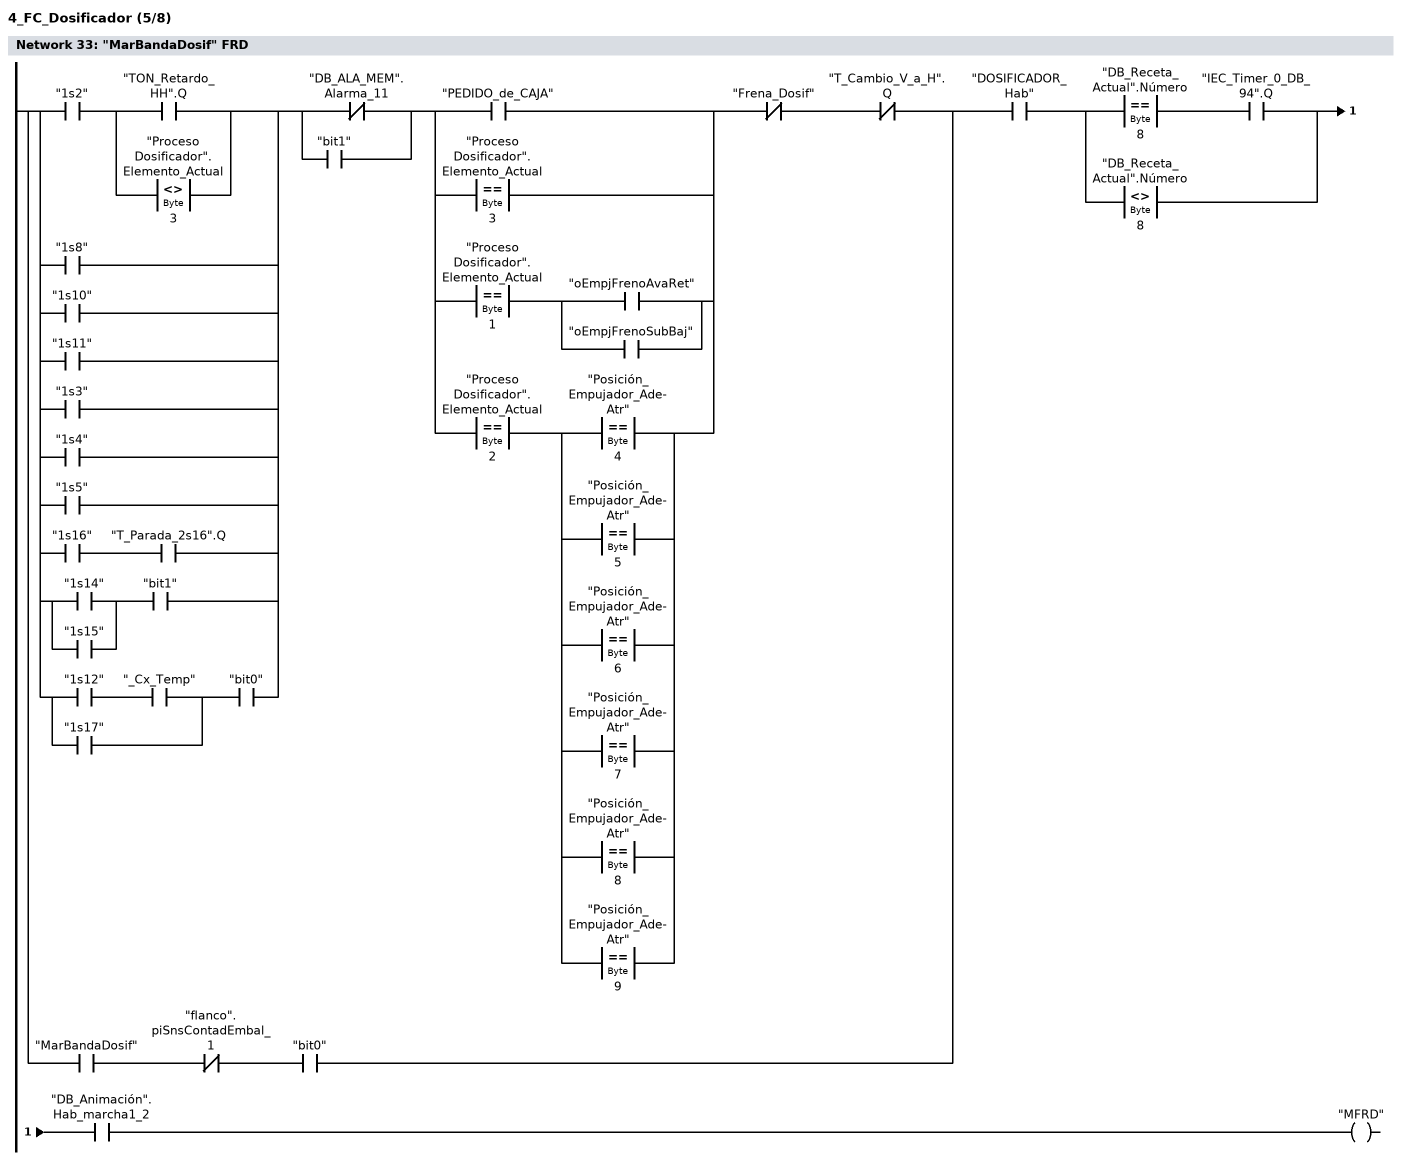
   RUNG wire#powerrail
      Contact( "1s2" )
      wire#w1
      Contact( "TON_Retardo_HH".Q )
      wire#w2
      I_Contact( "DB_ALA_MEM".Alarma_11 )
      wire#w5
      Contact( "PEDIDO_de_CAJA" )
      wire#w6
      I_Contact( "Frena_Dosif" )
      I_Contact( "T_Cambio_V_a_H".Q )
      wire#w9
      Contact( "DOSIFICADOR_Hab" )
      wire#w10
      { S7_Templates := "SrcType := Byte" } EQ_Contact(in1 := "DB_Receta_Actual".Número, in2 := 8)
      Contact( "IEC_Timer_0_DB_94".Q )
      wire#w11
      Contact( "DB_Animación".Hab_marcha1_2 )
      Coil( "MFRD" )
   END_RUNG
   RUNG wire#w1
      { S7_Templates := "SrcType := Byte" } NE_Contact(in1 := "Proceso Dosificador".Elemento_Actual, in2 := 3)
   END_RUNG wire#w2
   RUNG wire#powerrail
      Contact( "1s8" )
   END_RUNG wire#w2
   RUNG wire#powerrail
      Contact( "1s10" )
   END_RUNG wire#w2
   RUNG wire#powerrail
      Contact( "1s11" )
   END_RUNG wire#w2
   RUNG wire#powerrail
      Contact( "1s3" )
   END_RUNG wire#w2
   RUNG wire#powerrail
      Contact( "1s4" )
   END_RUNG wire#w2
   RUNG wire#powerrail
      Contact( "1s5" )
   END_RUNG wire#w2
   RUNG wire#powerrail
      Contact( "1s16" )
      Contact( "T_Parada_2s16".Q )
   END_RUNG wire#w2
   RUNG wire#powerrail
      Contact( "1s14" )
      wire#w3
      Contact( "bit1" )
   END_RUNG wire#w2
   RUNG wire#powerrail
      Contact( "1s15" )
   END_RUNG wire#w3
   RUNG wire#powerrail
      Contact( "1s12" )
      Contact( "_Cx_Temp" )
      wire#w4
      Contact( "bit0" )
   END_RUNG wire#w2
   RUNG wire#powerrail
      Contact( "1s17" )
   END_RUNG wire#w4
   RUNG wire#w2
      Contact( "bit1" )
   END_RUNG wire#w5
   RUNG wire#w5
      { S7_Templates := "SrcType := Byte" } EQ_Contact(in1 := "Proceso Dosificador".Elemento_Actual, in2 := 3)
   END_RUNG wire#w6
   RUNG wire#w5
      { S7_Templates := "SrcType := Byte" } EQ_Contact(in1 := "Proceso Dosificador".Elemento_Actual, in2 := 1)
      wire#w7
      Contact( "oEmpjFrenoAvaRet" )
   END_RUNG wire#w6
   RUNG wire#w7
      Contact( "oEmpjFrenoSubBaj" )
   END_RUNG wire#w6
   RUNG wire#w5
      { S7_Templates := "SrcType := Byte" } EQ_Contact(in1 := "Proceso Dosificador".Elemento_Actual, in2 := 2)
      wire#w8
      { S7_Templates := "SrcType := Byte" } EQ_Contact(in1 := "Posición_Empujador_Ade-Atr", in2 := 4)
   END_RUNG wire#w6
   RUNG wire#w8
      { S7_Templates := "SrcType := Byte" } EQ_Contact(in1 := "Posición_Empujador_Ade-Atr", in2 := 5)
   END_RUNG wire#w6
   RUNG wire#w8
      { S7_Templates := "SrcType := Byte" } EQ_Contact(in1 := "Posición_Empujador_Ade-Atr", in2 := 6)
   END_RUNG wire#w6
   RUNG wire#w8
      { S7_Templates := "SrcType := Byte" } EQ_Contact(in1 := "Posición_Empujador_Ade-Atr", in2 := 7)
   END_RUNG wire#w6
   RUNG wire#w8
      { S7_Templates := "SrcType := Byte" } EQ_Contact(in1 := "Posición_Empujador_Ade-Atr", in2 := 8)
   END_RUNG wire#w6
   RUNG wire#w8
      { S7_Templates := "SrcType := Byte" } EQ_Contact(in1 := "Posición_Empujador_Ade-Atr", in2 := 9)
   END_RUNG wire#w6
   RUNG wire#powerrail
      Contact( "MarBandaDosif" )
      I_Contact( "flanco".piSnsContadEmbal_1 )
      Contact( "bit0" )
   END_RUNG wire#w9
   RUNG wire#w10
      { S7_Templates := "SrcType := Byte" } NE_Contact(in1 := "DB_Receta_Actual".Número, in2 := 8)
   END_RUNG wire#w11
   // the same network as SCL:
   "MFRD" := (((("1s2" AND ("TON_Retardo_HH".Q OR ("Proceso Dosificador".Elemento_Actual <> 3))) OR "1s8" OR "1s10" OR "1s11" OR "1s3" OR "1s4" OR "1s5" OR ("1s16" AND "T_Parada_2s16".Q) OR (("1s14" OR "1s15") AND "bit1") OR ((("1s12" AND "_Cx_Temp") OR "1s17") AND "bit0")) AND (NOT "DB_ALA_MEM".Alarma_11 OR "bit1") AND ("PEDIDO_de_CAJA" OR ("Proceso Dosificador".Elemento_Actual = 3) OR (("Proceso Dosificador".Elemento_Actual = 1) AND ("oEmpjFrenoAvaRet" OR "oEmpjFrenoSubBaj")) OR (("Proceso Dosificador".Elemento_Actual = 2) AND (("Posición_Empujador_Ade-Atr" = 4) OR ("Posición_Empujador_Ade-Atr" = 5) OR ("Posición_Empujador_Ade-Atr" = 6) OR ("Posición_Empujador_Ade-Atr" = 7) OR ("Posición_Empujador_Ade-Atr" = 8) OR ("Posición_Empujador_Ade-Atr" = 9)))) AND NOT "Frena_Dosif" AND NOT "T_Cambio_V_a_H".Q) OR ("MarBandaDosif" AND NOT "flanco".piSnsContadEmbal_1 AND "bit0")) AND "DOSIFICADOR_Hab" AND ((("DB_Receta_Actual".Número = 8) AND "IEC_Timer_0_DB_94".Q) OR ("DB_Receta_Actual".Número <> 8)) AND "DB_Animación".Hab_marcha1_2;
END_REGION

REGION Network 34: "MarBandaDosif" IGS/CRJ
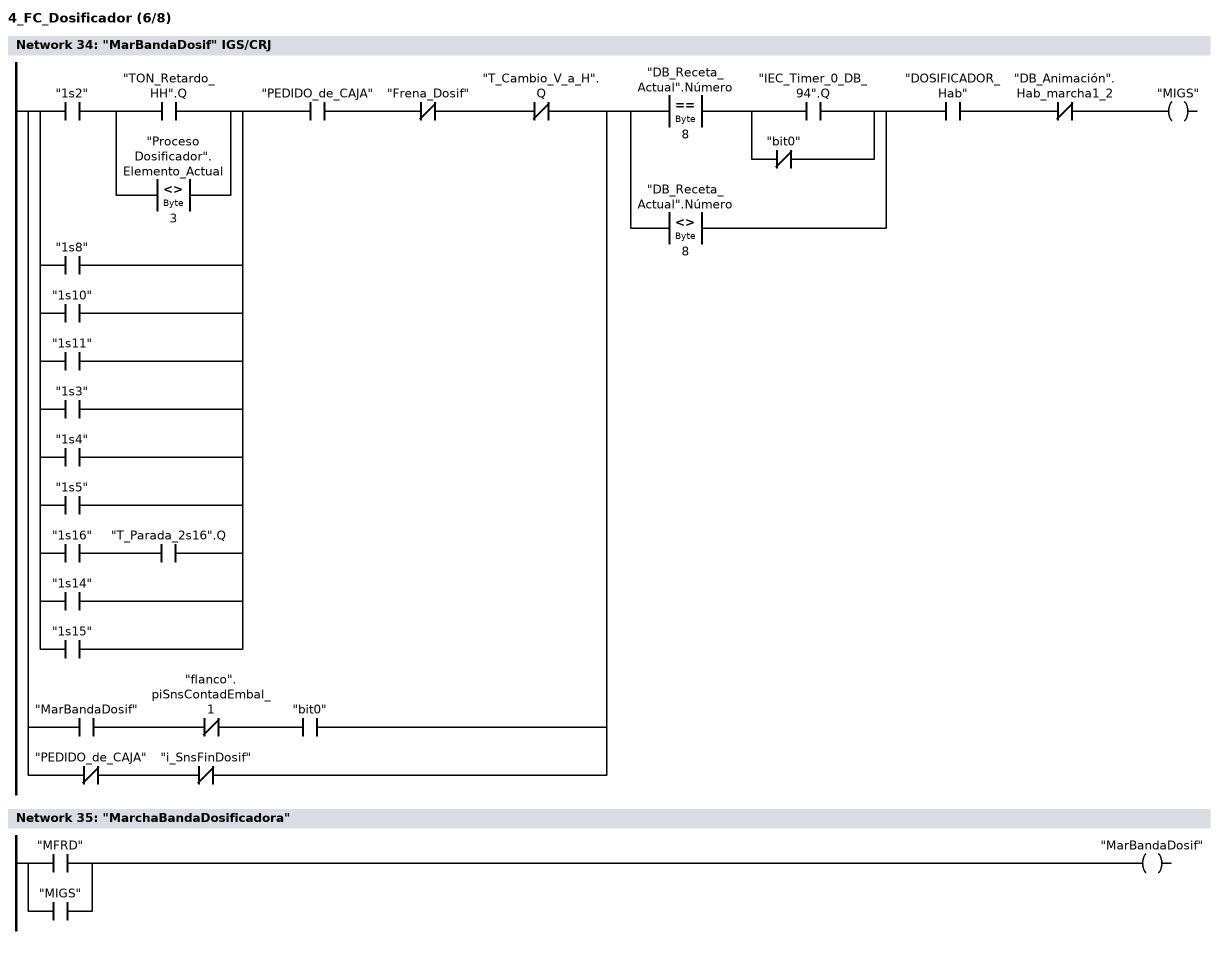
   RUNG wire#powerrail
      Contact( "1s2" )
      wire#w1
      Contact( "TON_Retardo_HH".Q )
      wire#w2
      Contact( "PEDIDO_de_CAJA" )
      I_Contact( "Frena_Dosif" )
      I_Contact( "T_Cambio_V_a_H".Q )
      wire#w3
      { S7_Templates := "SrcType := Byte" } EQ_Contact(in1 := "DB_Receta_Actual".Número, in2 := 8)
      wire#w4
      Contact( "IEC_Timer_0_DB_94".Q )
      wire#w5
      Contact( "DOSIFICADOR_Hab" )
      I_Contact( "DB_Animación".Hab_marcha1_2 )
      Coil( "MIGS" )
   END_RUNG
   RUNG wire#w1
      { S7_Templates := "SrcType := Byte" } NE_Contact(in1 := "Proceso Dosificador".Elemento_Actual, in2 := 3)
   END_RUNG wire#w2
   RUNG wire#powerrail
      Contact( "1s8" )
   END_RUNG wire#w2
   RUNG wire#powerrail
      Contact( "1s10" )
   END_RUNG wire#w2
   RUNG wire#powerrail
      Contact( "1s11" )
   END_RUNG wire#w2
   RUNG wire#powerrail
      Contact( "1s3" )
   END_RUNG wire#w2
   RUNG wire#powerrail
      Contact( "1s4" )
   END_RUNG wire#w2
   RUNG wire#powerrail
      Contact( "1s5" )
   END_RUNG wire#w2
   RUNG wire#powerrail
      Contact( "1s16" )
      Contact( "T_Parada_2s16".Q )
   END_RUNG wire#w2
   RUNG wire#powerrail
      Contact( "1s14" )
   END_RUNG wire#w2
   RUNG wire#powerrail
      Contact( "1s15" )
   END_RUNG wire#w2
   RUNG wire#powerrail
      Contact( "MarBandaDosif" )
      I_Contact( "flanco".piSnsContadEmbal_1 )
      Contact( "bit0" )
   END_RUNG wire#w3
   RUNG wire#powerrail
      I_Contact( "PEDIDO_de_CAJA" )
      I_Contact( "i_SnsFinDosif" )
   END_RUNG wire#w3
   RUNG wire#w4
      I_Contact( "bit0" )
   END_RUNG wire#w5
   RUNG wire#w3
      { S7_Templates := "SrcType := Byte" } NE_Contact(in1 := "DB_Receta_Actual".Número, in2 := 8)
   END_RUNG wire#w5
   // the same network as SCL:
   "MIGS" := (((("1s2" AND ("TON_Retardo_HH".Q OR ("Proceso Dosificador".Elemento_Actual <> 3))) OR "1s8" OR "1s10" OR "1s11" OR "1s3" OR "1s4" OR "1s5" OR ("1s16" AND "T_Parada_2s16".Q) OR "1s14" OR "1s15") AND "PEDIDO_de_CAJA" AND NOT "Frena_Dosif" AND NOT "T_Cambio_V_a_H".Q) OR ("MarBandaDosif" AND NOT "flanco".piSnsContadEmbal_1 AND "bit0") OR (NOT "PEDIDO_de_CAJA" AND NOT "i_SnsFinDosif")) AND ((("DB_Receta_Actual".Número = 8) AND ("IEC_Timer_0_DB_94".Q OR NOT "bit0")) OR ("DB_Receta_Actual".Número <> 8)) AND "DOSIFICADOR_Hab" AND NOT "DB_Animación".Hab_marcha1_2;
END_REGION

REGION Network 35: "MarchaBandaDosificadora"
   RUNG wire#powerrail
      Contact( "MFRD" )
      wire#w1
      Coil( "MarBandaDosif" )
   END_RUNG
   RUNG wire#powerrail
      Contact( "MIGS" )
   END_RUNG wire#w1
   // the same network as SCL:
   "MarBandaDosif" := "MFRD" OR "MIGS";
END_REGION

REGION Network 36: Temporizador provisario para Marcha Banda Dosifidicadora"
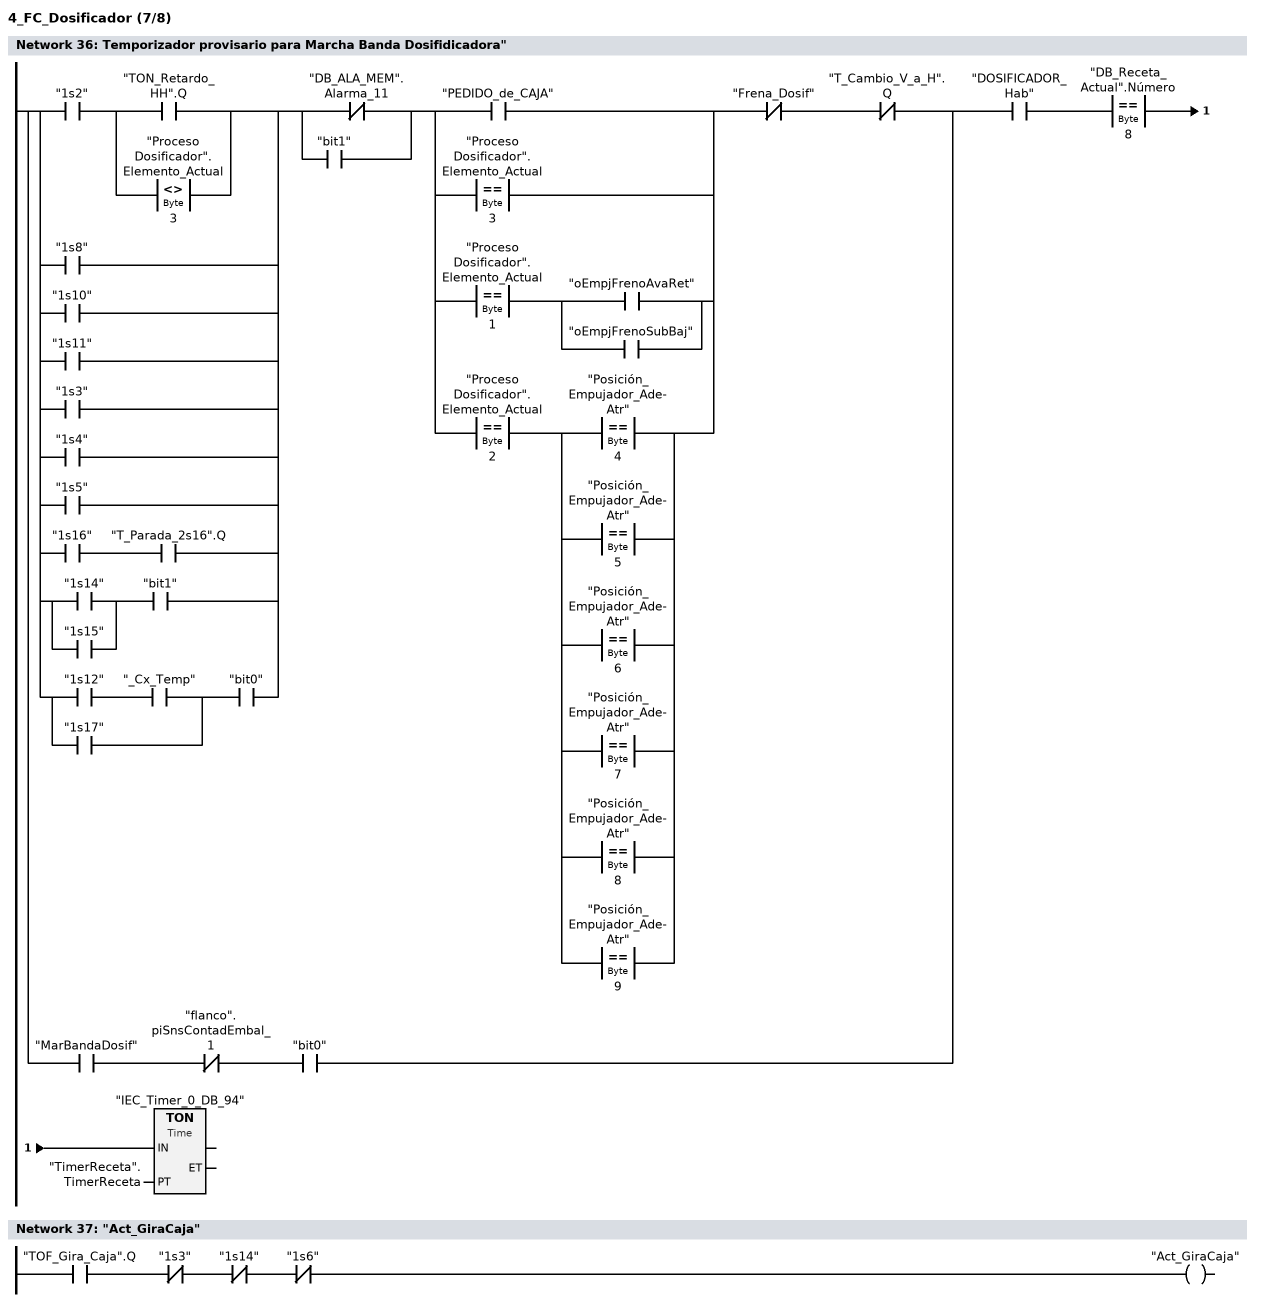
   "IEC_Timer_0_DB_94".TON(IN := (((("1s2" AND ("TON_Retardo_HH".Q OR ("Proceso Dosificador".Elemento_Actual <> 3))) OR "1s8" OR "1s10" OR "1s11" OR "1s3" OR "1s4" OR "1s5" OR ("1s16" AND "T_Parada_2s16".Q) OR (("1s14" OR "1s15") AND "bit1") OR ((("1s12" AND "_Cx_Temp") OR "1s17") AND "bit0")) AND (NOT "DB_ALA_MEM".Alarma_11 OR "bit1") AND ("PEDIDO_de_CAJA" OR ("Proceso Dosificador".Elemento_Actual = 3) OR (("Proceso Dosificador".Elemento_Actual = 1) AND ("oEmpjFrenoAvaRet" OR "oEmpjFrenoSubBaj")) OR (("Proceso Dosificador".Elemento_Actual = 2) AND (("Posición_Empujador_Ade-Atr" = 4) OR ("Posición_Empujador_Ade-Atr" = 5) OR ("Posición_Empujador_Ade-Atr" = 6) OR ("Posición_Empujador_Ade-Atr" = 7) OR ("Posición_Empujador_Ade-Atr" = 8) OR ("Posición_Empujador_Ade-Atr" = 9)))) AND NOT "Frena_Dosif" AND NOT "T_Cambio_V_a_H".Q) OR ("MarBandaDosif" AND NOT "flanco".piSnsContadEmbal_1 AND "bit0")) AND "DOSIFICADOR_Hab" AND ("DB_Receta_Actual".Número = 8),
                           PT := "TimerReceta".TimerReceta);
END_REGION

REGION Network 37: "Act_GiraCaja"
   RUNG wire#powerrail
      Contact( "TOF_Gira_Caja".Q )
      I_Contact( "1s3" )
      I_Contact( "1s14" )
      I_Contact( "1s6" )
      Coil( "Act_GiraCaja" )
   END_RUNG
   // the same network as SCL:
   "Act_GiraCaja" := "TOF_Gira_Caja".Q AND NOT "1s3" AND NOT "1s14" AND NOT "1s6";
END_REGION

REGION Network 38: "Act_EmpujaCaja"
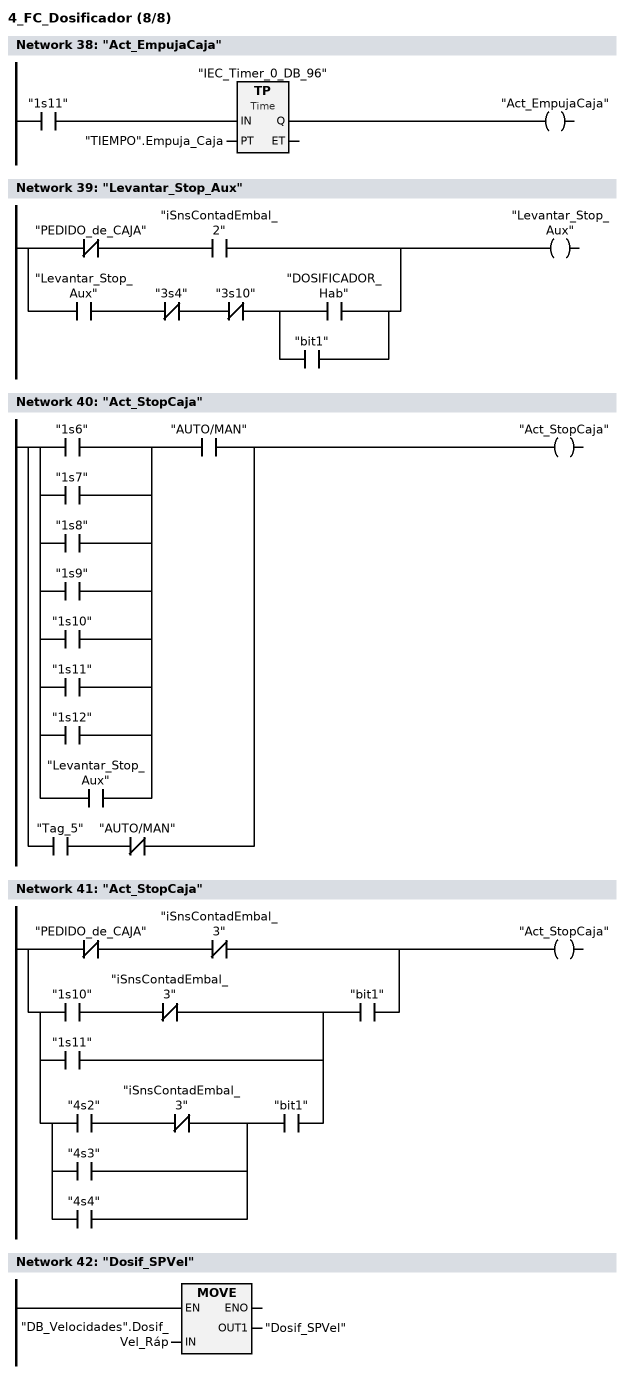
   "IEC_Timer_0_DB_96".TP(in := "1s11", pt := "TIEMPO".Empuja_Caja);
   "Act_EmpujaCaja" := "IEC_Timer_0_DB_96".q;
END_REGION

REGION Network 39: "Levantar_Stop_Aux"
   RUNG wire#powerrail
      I_Contact( "PEDIDO_de_CAJA" )
      Contact( "iSnsContadEmbal_2" )
      wire#w1
      Coil( "Levantar_Stop_Aux" )
   END_RUNG
   RUNG wire#powerrail
      Contact( "Levantar_Stop_Aux" )
      I_Contact( "3s4" )
      I_Contact( "3s10" )
      wire#w2
      Contact( "DOSIFICADOR_Hab" )
   END_RUNG wire#w1
   RUNG wire#w2
      Contact( "bit1" )
   END_RUNG wire#w1
   // the same network as SCL:
   "Levantar_Stop_Aux" := (NOT "PEDIDO_de_CAJA" AND "iSnsContadEmbal_2") OR ("Levantar_Stop_Aux" AND NOT "3s4" AND NOT "3s10" AND ("DOSIFICADOR_Hab" OR "bit1"));
END_REGION

REGION Network 40: "Act_StopCaja"
   RUNG wire#powerrail
      Contact( "1s6" )
      wire#w1
      Contact( "AUTO/MAN" )
      wire#w2
      Coil( "Act_StopCaja" )
   END_RUNG
   RUNG wire#powerrail
      Contact( "1s7" )
   END_RUNG wire#w1
   RUNG wire#powerrail
      Contact( "1s8" )
   END_RUNG wire#w1
   RUNG wire#powerrail
      Contact( "1s9" )
   END_RUNG wire#w1
   RUNG wire#powerrail
      Contact( "1s10" )
   END_RUNG wire#w1
   RUNG wire#powerrail
      Contact( "1s11" )
   END_RUNG wire#w1
   RUNG wire#powerrail
      Contact( "1s12" )
   END_RUNG wire#w1
   RUNG wire#powerrail
      Contact( "Levantar_Stop_Aux" )
   END_RUNG wire#w1
   RUNG wire#powerrail
      Contact( "Tag_5" )
      I_Contact( "AUTO/MAN" )
   END_RUNG wire#w2
   // the same network as SCL:
   "Act_StopCaja" := (("1s6" OR "1s7" OR "1s8" OR "1s9" OR "1s10" OR "1s11" OR "1s12" OR "Levantar_Stop_Aux") AND "AUTO/MAN") OR ("Tag_5" AND NOT "AUTO/MAN");
END_REGION

REGION Network 41: "Act_StopCaja"
   RUNG wire#powerrail
      I_Contact( "PEDIDO_de_CAJA" )
      I_Contact( "iSnsContadEmbal_3" )
      wire#w1
      Coil( "Act_StopCaja" )
   END_RUNG
   RUNG wire#powerrail
      Contact( "1s10" )
      I_Contact( "iSnsContadEmbal_3" )
      wire#w2
      Contact( "bit1" )
   END_RUNG wire#w1
   RUNG wire#powerrail
      Contact( "1s11" )
   END_RUNG wire#w2
   RUNG wire#powerrail
      Contact( "4s2" )
      I_Contact( "iSnsContadEmbal_3" )
      wire#w3
      Contact( "bit1" )
   END_RUNG wire#w2
   RUNG wire#powerrail
      Contact( "4s3" )
   END_RUNG wire#w3
   RUNG wire#powerrail
      Contact( "4s4" )
   END_RUNG wire#w3
   // the same network as SCL:
   "Act_StopCaja" := (NOT "PEDIDO_de_CAJA" AND NOT "iSnsContadEmbal_3") OR ((("1s10" AND NOT "iSnsContadEmbal_3") OR "1s11" OR ((("4s2" AND NOT "iSnsContadEmbal_3") OR "4s3" OR "4s4") AND "bit1")) AND "bit1");
END_REGION

REGION Network 42: "Dosif_SPVel"
   RUNG wire#powerrail
      { S7_GenerateENO := "TRUE" } Move(in := "DB_Velocidades".Dosif_Vel_Ráp, out1 => "Dosif_SPVel")
   END_RUNG
   // the same network as SCL:
   "Dosif_SPVel" := "DB_Velocidades".Dosif_Vel_Ráp;
END_REGION
END_FUNCTION

FUNCTION "5_FC_Empujador" : Void   // FC12, LAD
{ S7_Optimized_Access := 'FALSE' }
VERSION : 0.1
BEGIN

REGION Network 1
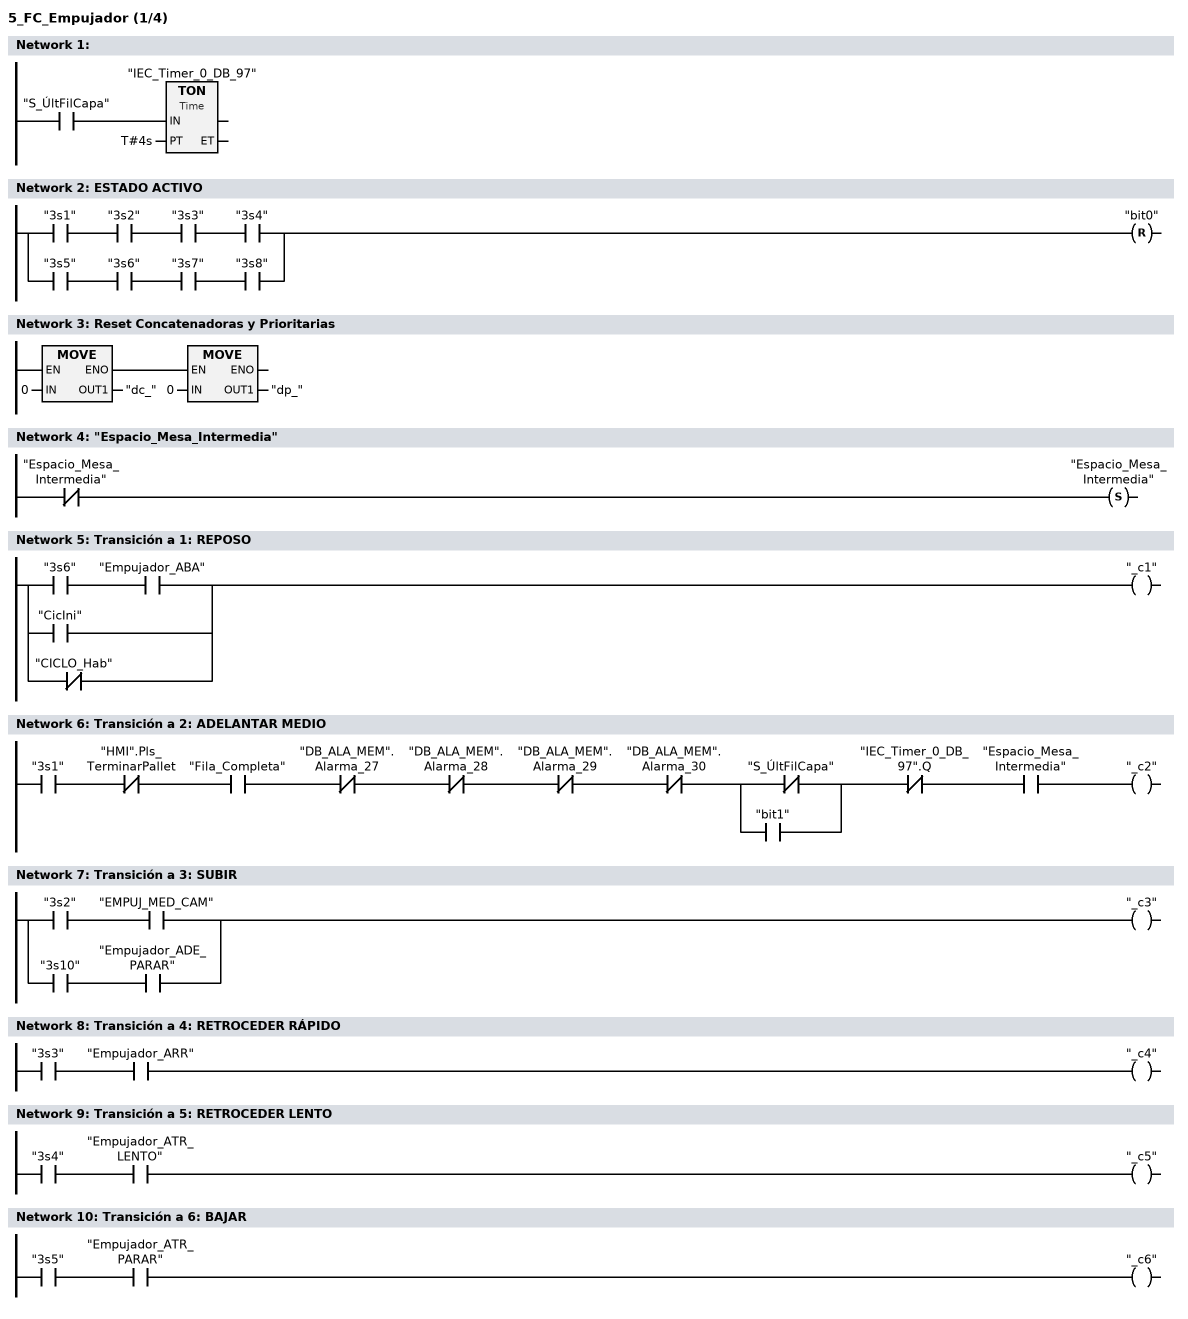
   "IEC_Timer_0_DB_97".TON(in := "S_ÚltFilCapa", pt := T#4s);
END_REGION

REGION Network 2: ESTADO ACTIVO
   RUNG wire#powerrail
      Contact( "3s1" )
      Contact( "3s2" )
      Contact( "3s3" )
      Contact( "3s4" )
      wire#w1
      R_Coil( "bit0" )
   END_RUNG
   RUNG wire#powerrail
      Contact( "3s5" )
      Contact( "3s6" )
      Contact( "3s7" )
      Contact( "3s8" )
   END_RUNG wire#w1
   // the same network as SCL:
   IF ("3s1" AND "3s2" AND "3s3" AND "3s4") OR ("3s5" AND "3s6" AND "3s7" AND "3s8") THEN
       "bit0" := FALSE;
   END_IF;
END_REGION

REGION Network 3: Reset Concatenadoras y Prioritarias
   RUNG wire#powerrail
      { S7_GenerateENO := "TRUE" } Move(in := 0, out1 => "dc_")
      { S7_GenerateENO := "TRUE" } Move(in := 0, out1 => "dp_")
   END_RUNG
   // the same network as SCL:
   // ENO of a box is taken as its EN; it also drops when the box reports an error
   "dc_" := 0;
   "dp_" := 0;
END_REGION

REGION Network 4: "Espacio_Mesa_Intermedia"
   RUNG wire#powerrail
      I_Contact( "Espacio_Mesa_Intermedia" )
      S_Coil( "Espacio_Mesa_Intermedia" )
   END_RUNG
   // the same network as SCL:
   IF NOT "Espacio_Mesa_Intermedia" THEN "Espacio_Mesa_Intermedia" := TRUE; END_IF;
END_REGION

REGION Network 5: Transición a 1: REPOSO
   RUNG wire#powerrail
      Contact( "3s6" )
      Contact( "Empujador_ABA" )
      wire#w1
      Coil( "_c1" )
   END_RUNG
   RUNG wire#powerrail
      Contact( "CicIni" )
   END_RUNG wire#w1
   RUNG wire#powerrail
      I_Contact( "CICLO_Hab" )
   END_RUNG wire#w1
   // the same network as SCL:
   "_c1" := ("3s6" AND "Empujador_ABA") OR "CicIni" OR NOT "CICLO_Hab";
END_REGION

REGION Network 6: Transición a 2: ADELANTAR MEDIO
   RUNG wire#powerrail
      Contact( "3s1" )
      I_Contact( "HMI".Pls_TerminarPallet )
      Contact( "Fila_Completa" )
      I_Contact( "DB_ALA_MEM".Alarma_27 )
      I_Contact( "DB_ALA_MEM".Alarma_28 )
      I_Contact( "DB_ALA_MEM".Alarma_29 )
      I_Contact( "DB_ALA_MEM".Alarma_30 )
      wire#w1
      I_Contact( "S_ÚltFilCapa" )
      wire#w2
      I_Contact( "IEC_Timer_0_DB_97".Q )
      Contact( "Espacio_Mesa_Intermedia" )
      Coil( "_c2" )
   END_RUNG
   RUNG wire#w1
      Contact( "bit1" )
   END_RUNG wire#w2
   // the same network as SCL:
   "_c2" := "3s1" AND NOT "HMI".Pls_TerminarPallet AND "Fila_Completa" AND NOT "DB_ALA_MEM".Alarma_27 AND NOT "DB_ALA_MEM".Alarma_28 AND NOT "DB_ALA_MEM".Alarma_29 AND NOT "DB_ALA_MEM".Alarma_30 AND (NOT "S_ÚltFilCapa" OR "bit1") AND NOT "IEC_Timer_0_DB_97".Q AND "Espacio_Mesa_Intermedia";
END_REGION

REGION Network 7: Transición a 3: SUBIR
   RUNG wire#powerrail
      Contact( "3s2" )
      Contact( "EMPUJ_MED_CAM" )
      wire#w1
      Coil( "_c3" )
   END_RUNG
   RUNG wire#powerrail
      Contact( "3s10" )
      Contact( "Empujador_ADE_PARAR" )
   END_RUNG wire#w1
   // the same network as SCL:
   "_c3" := ("3s2" AND "EMPUJ_MED_CAM") OR ("3s10" AND "Empujador_ADE_PARAR");
END_REGION

REGION Network 8: Transición a 4: RETROCEDER RÁPIDO
   RUNG wire#powerrail
      Contact( "3s3" )
      Contact( "Empujador_ARR" )
      Coil( "_c4" )
   END_RUNG
   // the same network as SCL:
   "_c4" := "3s3" AND "Empujador_ARR";
END_REGION

REGION Network 9: Transición a 5: RETROCEDER LENTO
   RUNG wire#powerrail
      Contact( "3s4" )
      Contact( "Empujador_ATR_LENTO" )
      Coil( "_c5" )
   END_RUNG
   // the same network as SCL:
   "_c5" := "3s4" AND "Empujador_ATR_LENTO";
END_REGION

REGION Network 10: Transición a 6: BAJAR
   RUNG wire#powerrail
      Contact( "3s5" )
      Contact( "Empujador_ATR_PARAR" )
      Coil( "_c6" )
   END_RUNG
   // the same network as SCL:
   "_c6" := "3s5" AND "Empujador_ATR_PARAR";
END_REGION

REGION Network 11: Transición a 7: ESPERAR PLATAFORMA
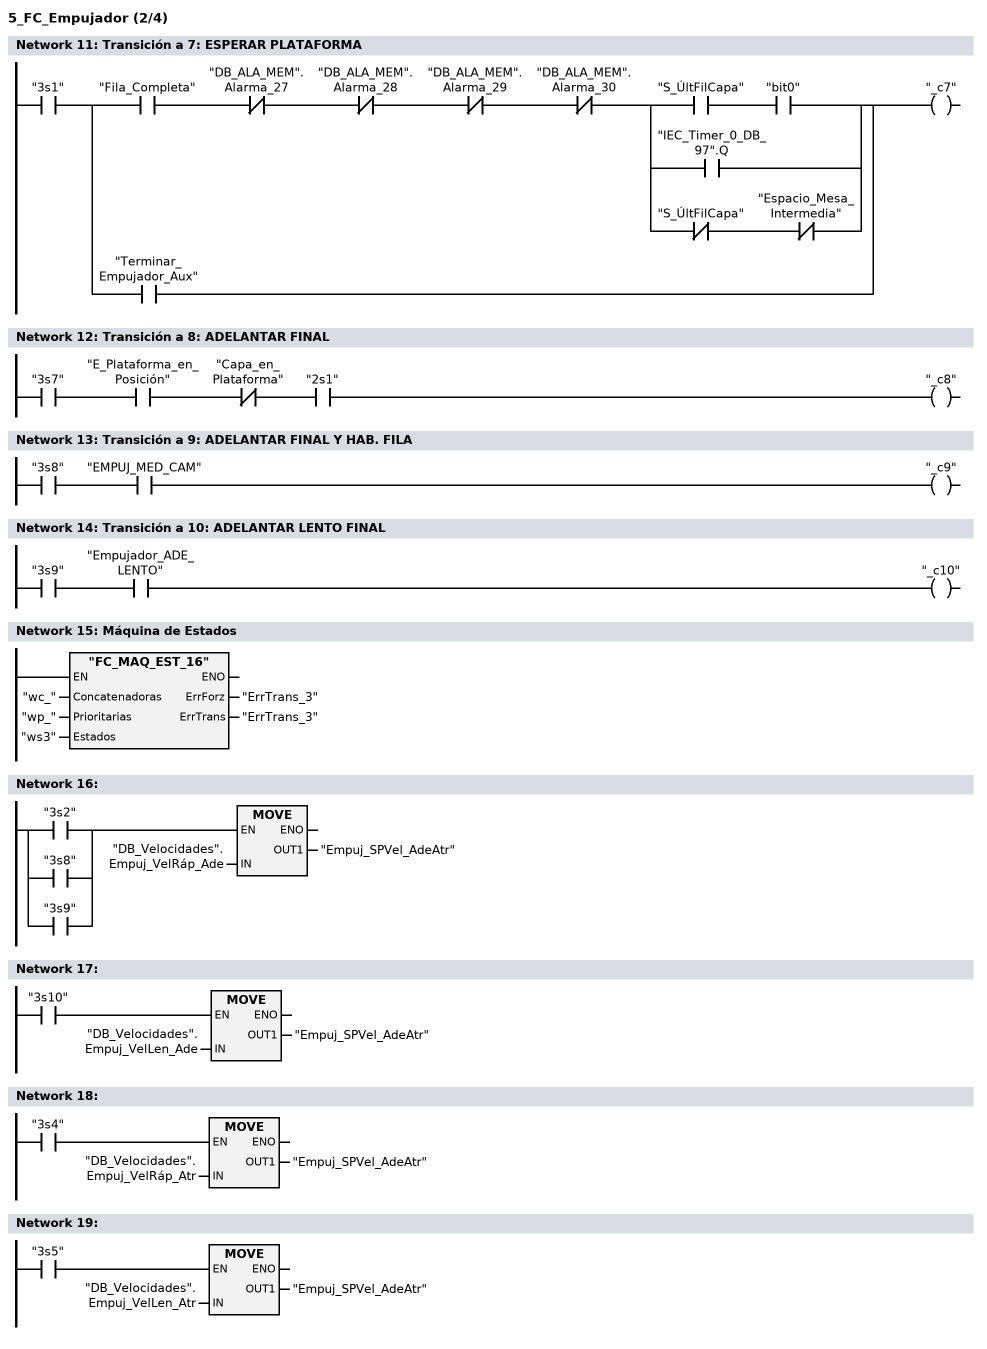
   RUNG wire#powerrail
      Contact( "3s1" )
      wire#w1
      Contact( "Fila_Completa" )
      I_Contact( "DB_ALA_MEM".Alarma_27 )
      I_Contact( "DB_ALA_MEM".Alarma_28 )
      I_Contact( "DB_ALA_MEM".Alarma_29 )
      I_Contact( "DB_ALA_MEM".Alarma_30 )
      wire#w2
      Contact( "S_ÚltFilCapa" )
      Contact( "bit0" )
      wire#w3
      Coil( "_c7" )
   END_RUNG
   RUNG wire#w2
      Contact( "IEC_Timer_0_DB_97".Q )
   END_RUNG wire#w3
   RUNG wire#w2
      I_Contact( "S_ÚltFilCapa" )
      I_Contact( "Espacio_Mesa_Intermedia" )
   END_RUNG wire#w3
   RUNG wire#w1
      Contact( "Terminar_Empujador_Aux" )
   END_RUNG wire#w3
   // the same network as SCL:
   "_c7" := "3s1" AND (("Fila_Completa" AND NOT "DB_ALA_MEM".Alarma_27 AND NOT "DB_ALA_MEM".Alarma_28 AND NOT "DB_ALA_MEM".Alarma_29 AND NOT "DB_ALA_MEM".Alarma_30 AND (("S_ÚltFilCapa" AND "bit0") OR "IEC_Timer_0_DB_97".Q OR (NOT "S_ÚltFilCapa" AND NOT "Espacio_Mesa_Intermedia"))) OR "Terminar_Empujador_Aux");
END_REGION

REGION Network 12: Transición a 8: ADELANTAR FINAL
   RUNG wire#powerrail
      Contact( "3s7" )
      Contact( "E_Plataforma_en_Posición" )
      I_Contact( "Capa_en_Plataforma" )
      Contact( "2s1" )
      Coil( "_c8" )
   END_RUNG
   // the same network as SCL:
   "_c8" := "3s7" AND "E_Plataforma_en_Posición" AND NOT "Capa_en_Plataforma" AND "2s1";
END_REGION

REGION Network 13: Transición a 9: ADELANTAR FINAL Y HAB. FILA
   RUNG wire#powerrail
      Contact( "3s8" )
      Contact( "EMPUJ_MED_CAM" )
      Coil( "_c9" )
   END_RUNG
   // the same network as SCL:
   "_c9" := "3s8" AND "EMPUJ_MED_CAM";
END_REGION

REGION Network 14: Transición a 10: ADELANTAR LENTO FINAL
   RUNG wire#powerrail
      Contact( "3s9" )
      Contact( "Empujador_ADE_LENTO" )
      Coil( "_c10" )
   END_RUNG
   // the same network as SCL:
   "_c10" := "3s9" AND "Empujador_ADE_LENTO";
END_REGION

REGION Network 15: Máquina de Estados
   RUNG wire#powerrail
      "FC_MAQ_EST_16"(Concatenadoras := "wc_", Prioritarias := "wp_", Estados := "ws3", ErrForz => "ErrTrans_3", ErrTrans => "ErrTrans_3")
   END_RUNG
   // the same network as SCL:
   "FC_MAQ_EST_16"(Concatenadoras := "wc_",
                   Prioritarias := "wp_",
                   Estados := "ws3",
                   ErrForz => "ErrTrans_3",
                   ErrTrans => "ErrTrans_3");
END_REGION

REGION Network 16
   RUNG wire#powerrail
      Contact( "3s2" )
      wire#w1
      { S7_GenerateENO := "TRUE" } Move(in := "DB_Velocidades".Empuj_VelRáp_Ade, out1 => "Empuj_SPVel_AdeAtr")
   END_RUNG
   RUNG wire#powerrail
      Contact( "3s8" )
   END_RUNG wire#w1
   RUNG wire#powerrail
      Contact( "3s9" )
   END_RUNG wire#w1
   // the same network as SCL:
   IF "3s2" OR "3s8" OR "3s9" THEN "Empuj_SPVel_AdeAtr" := "DB_Velocidades".Empuj_VelRáp_Ade; END_IF;
END_REGION

REGION Network 17
   RUNG wire#powerrail
      Contact( "3s10" )
      { S7_GenerateENO := "TRUE" } Move(in := "DB_Velocidades".Empuj_VelLen_Ade, out1 => "Empuj_SPVel_AdeAtr")
   END_RUNG
   // the same network as SCL:
   IF "3s10" THEN "Empuj_SPVel_AdeAtr" := "DB_Velocidades".Empuj_VelLen_Ade; END_IF;
END_REGION

REGION Network 18
   RUNG wire#powerrail
      Contact( "3s4" )
      { S7_GenerateENO := "TRUE" } Move(in := "DB_Velocidades".Empuj_VelRáp_Atr, out1 => "Empuj_SPVel_AdeAtr")
   END_RUNG
   // the same network as SCL:
   IF "3s4" THEN "Empuj_SPVel_AdeAtr" := "DB_Velocidades".Empuj_VelRáp_Atr; END_IF;
END_REGION

REGION Network 19
   RUNG wire#powerrail
      Contact( "3s5" )
      { S7_GenerateENO := "TRUE" } Move(in := "DB_Velocidades".Empuj_VelLen_Atr, out1 => "Empuj_SPVel_AdeAtr")
   END_RUNG
   // the same network as SCL:
   IF "3s5" THEN "Empuj_SPVel_AdeAtr" := "DB_Velocidades".Empuj_VelLen_Atr; END_IF;
END_REGION

REGION Network 20
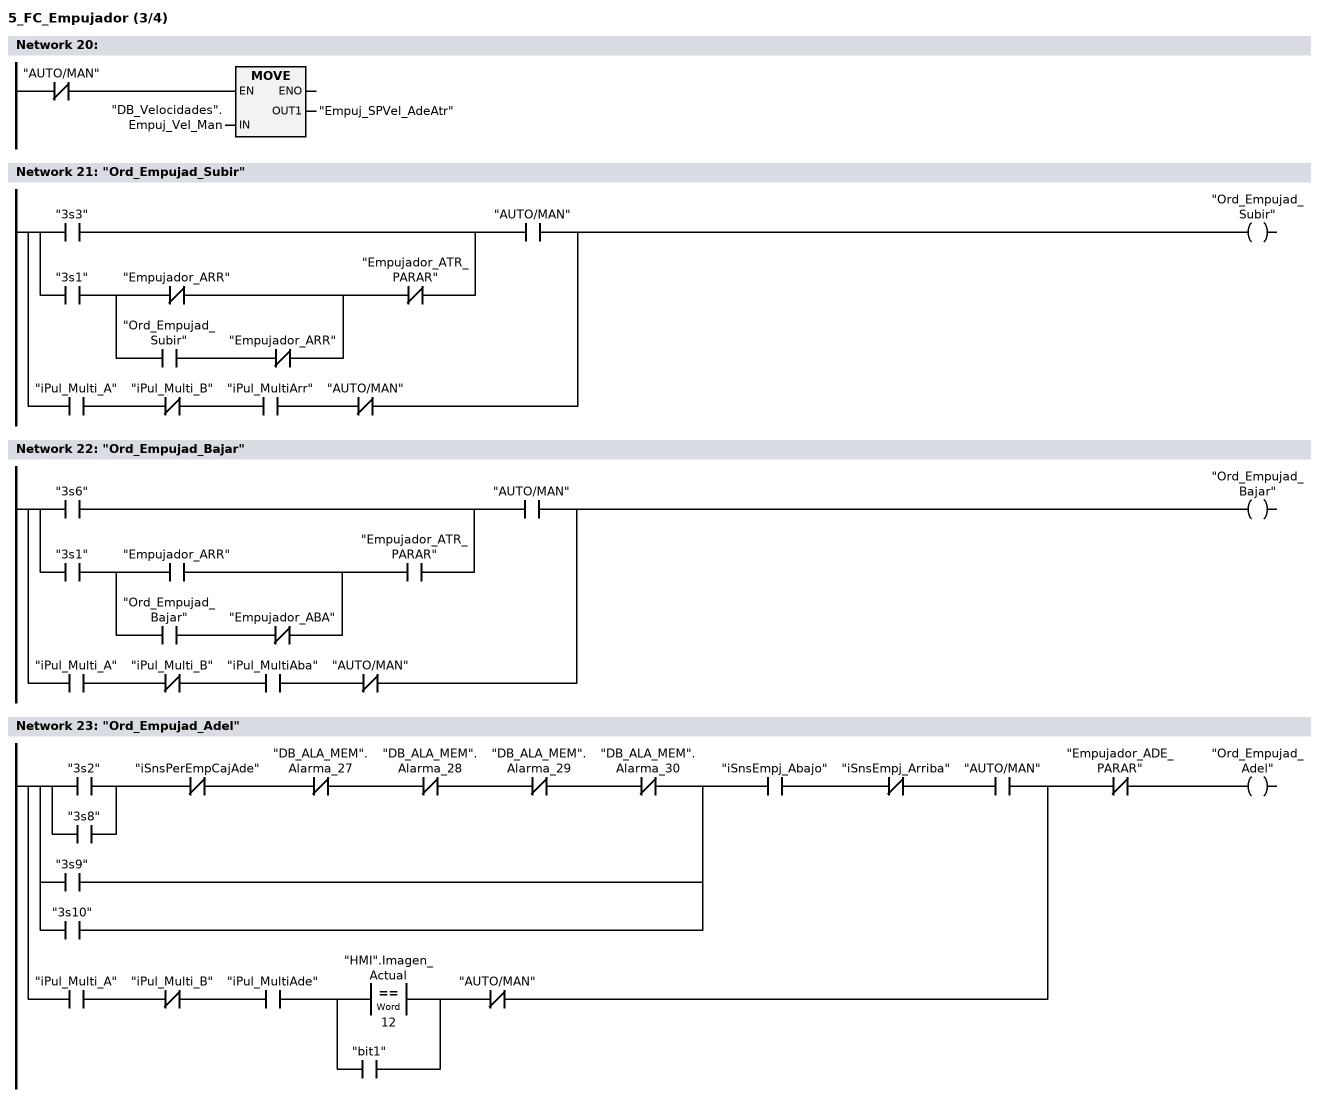
   RUNG wire#powerrail
      I_Contact( "AUTO/MAN" )
      { S7_GenerateENO := "TRUE" } Move(in := "DB_Velocidades".Empuj_Vel_Man, out1 => "Empuj_SPVel_AdeAtr")
   END_RUNG
   // the same network as SCL:
   IF NOT "AUTO/MAN" THEN "Empuj_SPVel_AdeAtr" := "DB_Velocidades".Empuj_Vel_Man; END_IF;
END_REGION

REGION Network 21: "Ord_Empujad_Subir"
   RUNG wire#powerrail
      Contact( "3s3" )
      wire#w1
      Contact( "AUTO/MAN" )
      wire#w4
      Coil( "Ord_Empujad_Subir" )
   END_RUNG
   RUNG wire#powerrail
      Contact( "3s1" )
      wire#w2
      I_Contact( "Empujador_ARR" )
      wire#w3
      I_Contact( "Empujador_ATR_PARAR" )
   END_RUNG wire#w1
   RUNG wire#w2
      Contact( "Ord_Empujad_Subir" )
      I_Contact( "Empujador_ARR" )
   END_RUNG wire#w3
   RUNG wire#powerrail
      Contact( "iPul_Multi_A" )
      I_Contact( "iPul_Multi_B" )
      Contact( "iPul_MultiArr" )
      I_Contact( "AUTO/MAN" )
   END_RUNG wire#w4
   // the same network as SCL:
   "Ord_Empujad_Subir" := (("3s3" OR ("3s1" AND (NOT "Empujador_ARR" OR ("Ord_Empujad_Subir" AND NOT "Empujador_ARR")) AND NOT "Empujador_ATR_PARAR")) AND "AUTO/MAN") OR ("iPul_Multi_A" AND NOT "iPul_Multi_B" AND "iPul_MultiArr" AND NOT "AUTO/MAN");
END_REGION

REGION Network 22: "Ord_Empujad_Bajar"
   RUNG wire#powerrail
      Contact( "3s6" )
      wire#w1
      Contact( "AUTO/MAN" )
      wire#w4
      Coil( "Ord_Empujad_Bajar" )
   END_RUNG
   RUNG wire#powerrail
      Contact( "3s1" )
      wire#w2
      Contact( "Empujador_ARR" )
      wire#w3
      Contact( "Empujador_ATR_PARAR" )
   END_RUNG wire#w1
   RUNG wire#w2
      Contact( "Ord_Empujad_Bajar" )
      I_Contact( "Empujador_ABA" )
   END_RUNG wire#w3
   RUNG wire#powerrail
      Contact( "iPul_Multi_A" )
      I_Contact( "iPul_Multi_B" )
      Contact( "iPul_MultiAba" )
      I_Contact( "AUTO/MAN" )
   END_RUNG wire#w4
   // the same network as SCL:
   "Ord_Empujad_Bajar" := (("3s6" OR ("3s1" AND ("Empujador_ARR" OR ("Ord_Empujad_Bajar" AND NOT "Empujador_ABA")) AND "Empujador_ATR_PARAR")) AND "AUTO/MAN") OR ("iPul_Multi_A" AND NOT "iPul_Multi_B" AND "iPul_MultiAba" AND NOT "AUTO/MAN");
END_REGION

REGION Network 23: "Ord_Empujad_Adel"
   RUNG wire#powerrail
      Contact( "3s2" )
      wire#w1
      I_Contact( "iSnsPerEmpCajAde" )
      I_Contact( "DB_ALA_MEM".Alarma_27 )
      I_Contact( "DB_ALA_MEM".Alarma_28 )
      I_Contact( "DB_ALA_MEM".Alarma_29 )
      I_Contact( "DB_ALA_MEM".Alarma_30 )
      wire#w2
      Contact( "iSnsEmpj_Abajo" )
      I_Contact( "iSnsEmpj_Arriba" )
      Contact( "AUTO/MAN" )
      wire#w3
      I_Contact( "Empujador_ADE_PARAR" )
      Coil( "Ord_Empujad_Adel" )
   END_RUNG
   RUNG wire#powerrail
      Contact( "3s8" )
   END_RUNG wire#w1
   RUNG wire#powerrail
      Contact( "3s9" )
   END_RUNG wire#w2
   RUNG wire#powerrail
      Contact( "3s10" )
   END_RUNG wire#w2
   RUNG wire#powerrail
      Contact( "iPul_Multi_A" )
      I_Contact( "iPul_Multi_B" )
      Contact( "iPul_MultiAde" )
      wire#w4
      { S7_Templates := "SrcType := Word" } EQ_Contact(in1 := "HMI".Imagen_Actual, in2 := 12)
      wire#w5
      I_Contact( "AUTO/MAN" )
   END_RUNG wire#w3
   RUNG wire#w4
      Contact( "bit1" )
   END_RUNG wire#w5
   // the same network as SCL:
   "Ord_Empujad_Adel" := ((((("3s2" OR "3s8") AND NOT "iSnsPerEmpCajAde" AND NOT "DB_ALA_MEM".Alarma_27 AND NOT "DB_ALA_MEM".Alarma_28 AND NOT "DB_ALA_MEM".Alarma_29 AND NOT "DB_ALA_MEM".Alarma_30) OR "3s9" OR "3s10") AND "iSnsEmpj_Abajo" AND NOT "iSnsEmpj_Arriba" AND "AUTO/MAN") OR ("iPul_Multi_A" AND NOT "iPul_Multi_B" AND "iPul_MultiAde" AND (("HMI".Imagen_Actual = 12) OR "bit1") AND NOT "AUTO/MAN")) AND NOT "Empujador_ADE_PARAR";
END_REGION

REGION Network 24: "Ord_Empujad_Atr"
